screen "05_Connection_Parameters" 800x480, template "Navigation"
   on GenerateScreen: SetTag("screen_number", 5)
   ScreenModuleView "Connection_Parameters_Control_1" at 100,137 size 600x270; ScreenModuleType ""
      on Guid_{11997190-31118}: ActivateScreen("03_Connection_Control", 0)
      Guid_{11997190-30476} <- "connection_parameters"
   Rectangle "screen_background" at 0,65 size 800x415
      Appearance <- "color"
      Visibility <- "visible"
*)

(* ===== HMI "HMI_RT_1" =====
system functions are stored by id; their names below are inferred from use

ScreenModuleEditorView "Row_Wire" 400x50
   Rectangle "Border" at 0,0 size 400x50
      Appearance <- "interface.background_animate"
   IOField "IOF R0 C0" at 5,5 size 190x45; FormatPattern ????????????????????
      ProcessValue <- "text_label"
      Appearance <- "interface.cell_0_animate"
      ObjectEnable <- "interface.cell_0_enable"
      Visibility <- "interface.cell_0_visible"
   IOField "IOF R0 C1" at 200,5 size 195x45; FormatPattern 9999999
      on OnFinishInput: SetBit("interface.cell_1_input_finished")
      Visibility <- "interface.cell_1_visible"
      ObjectEnable <- "interface.cell_1_enable"
      Appearance <- "interface.cell_1_animate"
*)

(* ===== HMI "HMI_RT_1" =====
system functions are stored by id; their names below are inferred from use

ScreenModuleEditorView "Row_Wire" 400x50
   Rectangle "Border" at 0,0 size 400x50
      Appearance <- "interface.background_animate"
      Visibility <- "interface.background_visible"
   IOField "IOF R0 C0" at 5,5 size 190x45; FormatPattern ????????????????????
      Appearance <- "interface.cell_0_animate"
      ProcessValue <- "text_label"
      Visibility <- "interface.cell_0_visible"
      ObjectEnable <- "interface.cell_0_enable"
   IOField "IOF R0 C1" at 200,5 size 195x45; FormatPattern 9999999
      on OnFinishInput: SetBit("interface.cell_1_input_finished")
      Visibility <- "interface.cell_1_visible"
      Appearance <- "interface.cell_1_animate"
      ObjectEnable <- "interface.cell_1_enable"
*)

(* ===== HMI "HMI_RT_1" =====
system functions are stored by id; their names below are inferred from use

ScreenModuleEditorView "Row_Wire" 400x50
   Rectangle "Border" at 0,0 size 400x50
      Visibility <- "interface.background_visible"
      Appearance <- "interface.background_animate"
   IOField "IOF R0 C0" at 5,5 size 190x45; FormatPattern ????????????????????
      Appearance <- "interface.cell_0_animate"
      Visibility <- "interface.cell_0_visible"
      ObjectEnable <- "interface.cell_0_enable"
      ProcessValue <- "interface.cell_0_value"
   IOField "IOF R0 C1" at 200,5 size 195x45; FormatPattern 9999999
      on OnFinishInput: SetBit("interface.cell_1_input_finished")
      Visibility <- "interface.cell_1_visible"
      Appearance <- "interface.cell_1_animate"
      ObjectEnable <- "interface.cell_1_enable"
*)

(* ===== HMI "HMI_RT_1" =====
system functions are stored by id; their names below are inferred from use

ScreenModuleEditorView "Row_Wire" 400x50
   Rectangle "Border" at 0,0 size 400x50
      Visibility <- "interface.background_visible"
      Appearance <- "interface.background_animate"
   IOField "IOF R0 C0" at 5,5 size 190x45; FormatPattern ????????????????????
      Appearance <- "interface.cell_0_animate"
      Visibility <- "interface.cell_0_visible"
      ProcessValue <- "interface.cell_0_value"
      ObjectEnable <- "interface.cell_0_enable"
   IOField "IOF R0 C1" at 200,5 size 195x45; FormatPattern 9999999
      on OnFinishInput: SetBit("interface.cell_1_input_finished")
      Visibility <- "interface.cell_1_visible"
      Appearance <- "interface.cell_1_animate"
      ObjectEnable <- "interface.cell_1_enable"
*)

(* ===== HMI "HMI_RT_1" =====
system functions are stored by id; their names below are inferred from use

ScreenModuleEditorView "Row_Wire" 400x65
   Rectangle "Border" at 0,0 size 400x65
      Visibility <- "interface.background_visible"
      Appearance <- "interface.background_animate"
   TextField "TF R0 C0" at 5,5 size 190x60; Text 'Text'
      Visibility <- "interface.cell_0_visible"
   IOField "IOF R0 C1" at 200,5 size 195x60; FormatPattern 9999999
      on OnFinishInput: SetBit("interface.cell_1_input_finished")
      Visibility <- "interface.cell_1_visible"
      ObjectEnable <- "interface.cell_1_enable"
*)

(* ===== HMI "HMI_RT_1" =====
system functions are stored by id; their names below are inferred from use

ScreenModuleEditorView "Row_Wire" 600x65
   Rectangle "Border" at 0,0 size 600x65
      Visibility <- "interface.background_visible"
      Appearance <- "interface.background_animate"
   TextField "TF R0 C0" at 5,5 size 360x60; Text 'CARBON WIRE'
      Visibility <- "interface.cell_0_visible"
   IOField "IOF R0 C1" at 370,5 size 225x60; FormatPattern 9999999
      on OnFinishInput: SetBit("interface.cell_1_input_finished")
      Visibility <- "interface.cell_1_visible"
      ObjectEnable <- "interface.cell_1_enable"
*)

(* ===== HMI "HMI_RT_1" =====
system functions are stored by id; their names below are inferred from use

ScreenModuleEditorView "Row_Wire" 600x65
   Rectangle "Border" at 0,0 size 600x65
      Visibility <- "interface.background_visible"
      Appearance <- "interface.background_animate"
   TextField "TF R0 C0" at 5,5 size 360x60; Text 'CARBON WIRE'
      Visibility <- "interface.cell_0_visible"
      Appearance <- "interface.cell_0_animate"
   IOField "IOF R0 C1" at 370,5 size 225x60; FormatPattern 9999999
      on OnFinishInput: SetBit("interface.cell_1_input_finished")
      Visibility <- "interface.cell_1_visible"
      ObjectEnable <- "interface.cell_1_enable"
      Appearance <- "interface.cell_1_animate"
*)

(* ===== HMI "HMI_RT_1" =====
system functions are stored by id; their names below are inferred from use

ScreenModuleEditorView "Row_Wire_Label" 600x65
   Rectangle "Border" at 0,0 size 600x65
      Visibility <- "interface.background_visible"
      Appearance <- "interface.background_animate"
   TextField "TF R0 C0" at 5,5 size 360x60; Text 'CARBON WIRE'
      Visibility <- "interface.cell_0_visible"
      Appearance <- "interface.cell_0_animate"
   IOField "IOF R0 C1" at 370,5 size 225x60; FormatPattern 9999999
      on OnFinishInput: SetBit("interface.cell_1_input_finished")
      Visibility <- "interface.cell_1_visible"
      Appearance <- "interface.cell_1_animate"
      ObjectEnable <- "interface.cell_1_enable"
*)

(* ===== HMI "HMI_RT_1" =====

ScreenModuleEditorView "Row_Wire_Label" 600x65
   Rectangle "Border" at 0,0 size 600x65
      Visibility <- "interface.background_visible"
      Appearance <- "interface.background_animate"
   TextField "TF R0 C0" at 5,5 size 360x60; Text 'WIRE'
      Visibility <- "interface.cell_0_visible"
      Appearance <- "interface.cell_0_animate"
   TextField "TF R0 C1" at 370,5 size 225x60; Text 'LENGTH'
      Visibility <- "interface.cell_1_visible"
      Appearance <- "interface.cell_1_animate"
*)

(* ===== HMI "HMI_RT_1" =====

ScreenModuleEditorView "Divider" 600x5
   Line "line" at 10,2 size 580x0
      Appearance <- "interface.line_animate"
      Visibility <- "interface.line_visible"
   Rectangle "background" at 0,0 size 600x5
      Appearance <- "interface.background_animate"
      Visibility <- "interface.background_visible"
*)

(* ===== HMI "HMI_RT_1" =====
system functions are stored by id; their names below are inferred from use

ScreenModuleEditorView "Navigation" 800x65
   Button "Wire" at 5,5 size 390x60; TextOff 'WIRE'
      Appearance <- "interface.wire_animate"
      on Press: function_b14e0dd5("interface.wire_actuate", 0)
   Button "Material" at 400,5 size 390x60; TextOff 'MATERIAL'
      Appearance <- "interface.material_animate"
      on Press: function_b14e0dd5("interface.material_actuate", 0)
   Rectangle "Wire_Cover" at 10,60 size 380x5
      Visibility <- "interface.wire_cover_visible"
   Rectangle "Material_Cover" at 405,60 size 380x5
      Visibility <- "interface.material_cover_visible"
*)

(* ===== HMI "HMI_RT_1" =====
system functions are stored by id; their names below are inferred from use

ScreenModuleEditorView "Navigation" 800x65
   Button "Wire" at 5,5 size 390x60; TextOff 'WIRE'
      on Press: function_b14e0dd5("interface.wire_actuate", 0)
      Appearance <- "interface.wire_animate"
   Button "Material" at 400,5 size 390x60; TextOff 'MATERIAL'
      on Press: function_b14e0dd5("interface.material_actuate", 0)
      Appearance <- "interface.material_animate"
   Rectangle "Wire_Cover" at 10,60 size 380x5
      Visibility <- "interface.wire_cover_visible"
   Rectangle "Material_Cover" at 405,60 size 380x5
      Visibility <- "interface.material_cover_visible"
*)

(* ===== HMI "HMI_RT_1" =====
system functions are stored by id; their names below are inferred from use

ScreenModuleEditorView "Navigation" 800x65
   Button "Wire" at 5,5 size 392x60; TextOff 'WIRE'
      on Press: function_b14e0dd5("interface.wire_actuate", 0)
      Appearance <- "interface.wire_animate"
   Button "Material" at 402,5 size 393x60; TextOff 'MATERIAL'
      on Press: function_b14e0dd5("interface.material_actuate", 0)
      Appearance <- "interface.material_animate"
   Rectangle "Wire_Cover" at 10,60 size 382x5
      Visibility <- "interface.wire_cover_visible"
   Rectangle "Material_Cover" at 407,60 size 383x5
      Visibility <- "interface.material_cover_visible"
*)

(* ===== HMI "HMI_RT_1" =====
system functions are stored by id; their names below are inferred from use

ScreenModuleEditorView "Row_Material" 600x65
   Rectangle "Border" at 0,0 size 600x65
      Visibility <- "interface.background_visible"
      Appearance <- "interface.background_animate"
   TextField "TF R0 C0" at 5,5 size 360x60; Text 'CARBON WIRE'
      Visibility <- "interface.cell_0_visible"
      Appearance <- "interface.cell_0_animate"
   IOField "IOF R0 C1" at 370,5 size 225x60; FormatPattern 9999999
      on OnFinishInput: SetBit("interface.cell_1_input_finished")
      Visibility <- "interface.cell_1_visible"
      Appearance <- "interface.cell_1_animate"
      ObjectEnable <- "interface.cell_1_enable"
*)

(* ===== HMI "HMI_RT_1" =====
system functions are stored by id; their names below are inferred from use

ScreenModuleEditorView "Row_Material" 600x40
   Rectangle "Border" at 0,0 size 600x40
      Visibility <- "interface.background_visible"
      Appearance <- "interface.background_animate"
   IOField "IOF R0 C1" at 370,5 size 225x35; FormatPattern 9999999
      on OnFinishInput: SetBit("interface.cell_1_input_finished")
      Visibility <- "interface.cell_1_visible"
      Appearance <- "interface.cell_1_animate"
      ObjectEnable <- "interface.cell_1_enable"
   TextField "TF R0 C0" at 5,5 size 360x35; Text 'MOLYBDENUM'
      Visibility <- "interface.cell_0_visible"
      Appearance <- "interface.cell_0_animate"
*)

(* ===== HMI "HMI_RT_1" =====
system functions are stored by id; their names below are inferred from use

ScreenModuleEditorView "Row_Custom" 600x40
   Rectangle "Border" at 0,0 size 600x40
      Visibility <- "interface.background_visible"
      Appearance <- "interface.background_animate"
   IOField "IOF R0 C1" at 370,5 size 225x35; FormatPattern 9999999
      on OnFinishInput: SetBit("interface.cell_1_input_finished")
      Visibility <- "interface.cell_1_visible"
      Appearance <- "interface.cell_1_animate"
      ObjectEnable <- "interface.cell_1_enable"
   TextField "TF R0 C0" at 5,5 size 360x35; Text 'MOLYBDENUM'
      Visibility <- "interface.cell_0_visible"
      Appearance <- "interface.cell_0_animate"
*)

(* ===== HMI "HMI_RT_1" =====
system functions are stored by id; their names below are inferred from use

ScreenModuleEditorView "Row_Custom" 600x40
   Rectangle "Border" at 0,0 size 600x40
      Visibility <- "interface.background_visible"
      Appearance <- "interface.background_animate"
   IOField "IOF R0 C0" at 5,5 size 360x35; FormatPattern ???????????????
      on OnFinishInput: SetBit("interface.cell_0_input_finished")
      Appearance <- "interface.cell_0_animate"
      ObjectEnable <- "interface.cell_0_enable"
      Visibility <- "interface.cell_0_visible"
   IOField "IOF R0 C1" at 370,5 size 225x35; FormatPattern 9999999
      on OnFinishInput: SetBit("interface.cell_1_input_finished")
      Visibility <- "interface.cell_1_visible"
      Appearance <- "interface.cell_1_animate"
      ObjectEnable <- "interface.cell_1_enable"
*)

(* ===== HMI "HMI_RT_1" =====
system functions are stored by id; their names below are inferred from use

ScreenModuleEditorView "Row_Material_Label" 600x40
   Rectangle "Border" at 0,0 size 600x40
      Visibility <- "interface.background_visible"
      Appearance <- "interface.background_animate"
   IOField "IOF R0 C1" at 370,5 size 225x35; FormatPattern 9999999
      on OnFinishInput: SetBit("interface.cell_1_input_finished")
      Visibility <- "interface.cell_1_visible"
      Appearance <- "interface.cell_1_animate"
      ObjectEnable <- "interface.cell_1_enable"
   TextField "TF R0 C0" at 5,5 size 360x35; Text 'MOLYBDENUM'
      Visibility <- "interface.cell_0_visible"
      Appearance <- "interface.cell_0_animate"
*)

(* ===== HMI "HMI_RT_1" =====

ScreenModuleEditorView "Row_Material_Label" 600x40
   Rectangle "Border" at 0,0 size 600x40
      Visibility <- "interface.background_visible"
      Appearance <- "interface.background_animate"
   TextField "TF R0 C0" at 5,5 size 360x35; Text 'MATERIAL'
      Visibility <- "interface.cell_0_visible"
      Appearance <- "interface.cell_0_animate"
   TextField "TF R0 C1" at 370,5 size 225x35; Text 'BAGS'
      Appearance <- "interface.cell_1_animate"
      Visibility <- "interface.cell_1_visible"
*)

(* ===== HMI "HMI_RT_1" =====
system functions are stored by id; their names below are inferred from use

ScreenModuleEditorView "Row_Wire" 600x65
   Rectangle "Border" at 0,0 size 600x65
      Visibility <- "interface.background_visible"
   TextField "TF R0 C0" at 5,5 size 360x60; Text 'CARBON WIRE'
      Visibility <- "interface.cell_0_visible"
   IOField "IOF R0 C1" at 370,5 size 225x60; FormatPattern 9999999
      on OnFinishInput: SetBit("interface.cell_1_input_finished")
      Visibility <- "interface.cell_1_visible"
      Appearance <- "interface.cell_1_animate"
      ObjectEnable <- "interface.cell_1_enable"
      on Activate: SetBit("interface.cell_1_active")
      on Deactivate: ResetBit("interface.cell_1_active")
*)

(* ===== HMI "HMI_RT_1" =====

ScreenModuleEditorView "Divider" 600x5
   Line "line" at 10,2 size 580x0
      Visibility <- "interface.line_visible"
      Appearance <- "interface.line_animate"
   Rectangle "background" at 0,0 size 600x5
      Visibility <- "interface.background_visible"
      Appearance <- "interface.background_animate"
*)

(* ===== HMI "HMI_RT_1" =====
system functions are stored by id; their names below are inferred from use

ScreenModuleEditorView "Row_Material" 600x40
   Rectangle "Border" at 0,0 size 600x40
      Visibility <- "interface.background_visible"
      Appearance <- "interface.background_animate"
   IOField "IOF R0 C1" at 370,5 size 225x35; FormatPattern 9999999
      on OnFinishInput: SetBit("interface.cell_1_input_finished")
      Visibility <- "interface.cell_1_visible"
      Appearance <- "interface.cell_1_animate"
      ObjectEnable <- "interface.cell_1_enable"
   TextField "TF R0 C0" at 5,5 size 360x35; Text 'MOLYBDENUM'
      Visibility <- "interface.cell_0_visible"
      Appearance <- "interface.cell_0_animate"
*)

(* ===== HMI "HMI_RT_1" =====
system functions are stored by id; their names below are inferred from use

ScreenModuleEditorView "Navigation" 800x65
   Button "Wire" at 5,5 size 392x60; TextOff 'WIRE'
      on Press: function_b14e0dd5("interface.wire_actuate", 0)
      Appearance <- "interface.wire_animate"
      ObjectEnable <- "interface.wire_enable"
      Visibility <- "interface.wire_visible"
   Button "Material" at 402,5 size 393x60; TextOff 'MATERIAL'
      on Press: function_b14e0dd5("interface.material_actuate", 0)
      Appearance <- "interface.material_animate"
      ObjectEnable <- "interface.material_enable"
      Visibility <- "interface.material_visible"
   Rectangle "Background" at 0,0 size 800x65
      Appearance <- "interface.background_animate"
      Visibility <- "interface.background_visible"
   Rectangle "Wire_Cover" at 10,60 size 382x5
      Visibility <- "interface.wire_cover_visible"
      Appearance <- "interface.wire_cover_animate"
   Rectangle "Material_Cover" at 407,60 size 383x5
      Visibility <- "interface.material_cover_visible"
      Appearance <- "interface.material_cover_animate"
   Line "Bottom_Line" at 0,62 size 800x0
      Appearance <- "interface.bottom_line_animate"
      Visibility <- "interface.bottom_line_visible"
*)

(* ===== HMI "HMI_RT_1" =====
system functions are stored by id; their names below are inferred from use

ScreenModuleEditorView "Navigation" 800x65
   Button "Wire" at 5,5 size 392x60; TextOff 'WIRE'
      on Press: function_b14e0dd5("interface.wire_actuate", 0)
      Appearance <- "interface.wire_animate"
      ObjectEnable <- "interface.wire_enable"
      Visibility <- "interface.wire_visible"
   Button "Material" at 402,5 size 393x60; TextOff 'MATERIAL'
      on Press: function_b14e0dd5("interface.material_actuate", 0)
      Appearance <- "interface.material_animate"
      ObjectEnable <- "interface.material_enable"
      Visibility <- "interface.material_visible"
   Rectangle "Background" at 0,0 size 800x65
      Visibility <- "interface.background_visible"
      Appearance <- "interface.background_animate"
   Rectangle "Wire_Cover" at 10,60 size 382x5
      Visibility <- "interface.wire_cover_visible"
      Appearance <- "interface.wire_cover_animate"
   Rectangle "Material_Cover" at 407,60 size 383x5
      Visibility <- "interface.material_cover_visible"
      Appearance <- "interface.material_cover_animate"
   Line "Bottom_Line" at 0,62 size 800x0
      Visibility <- "interface.bottom_line_visible"
      Appearance <- "interface.bottom_line_animate"
*)

(* ===== HMI "HMI_RT_1" =====
system functions are stored by id; their names below are inferred from use

ScreenModuleEditorView "Navigation" 800x65
   Button "Wire" at 5,5 size 392x60; TextOff 'WIRE'
      on Press: function_b14e0dd5("interface.wire_actuate", 0)
      Appearance <- "interface.wire_animate"
      ObjectEnable <- "interface.wire_enable"
      Visibility <- "interface.wire_visible"
   Button "Material" at 402,5 size 393x60; TextOff 'MATERIAL'
      on Press: function_b14e0dd5("interface.material_actuate", 0)
      Appearance <- "interface.material_animate"
      ObjectEnable <- "interface.material_enable"
      Visibility <- "interface.material_visible"
   Rectangle "Background" at 0,0 size 800x65
      Visibility <- "interface.background_visible"
      Appearance <- "interface.background_animate"
   Rectangle "Wire_Cover" at 10,60 size 382x5
      Visibility <- "interface.wire_cover_visible"
      Appearance <- "interface.wire_cover_animate"
   Rectangle "Material_Cover" at 407,60 size 383x5
      Visibility <- "interface.material_cover_visible"
      Appearance <- "interface.material_cover_animate"
   Line "Bottom_Line" at 0,62 size 800x0
      Visibility <- "interface.bottom_line_visible"
      Appearance <- "interface.bottom_line_animate"
*)

(* ===== HMI "HMI_RT_1" =====
system functions are stored by id; their names below are inferred from use

ScreenModuleEditorView "Navigation" 800x65
   Button "Wire" at 5,5 size 392x60; TextOff 'WIRE'
      on Press: function_b14e0dd5("interface.wire_actuate", 0)
      Appearance <- "interface.wire_animate"
      ObjectEnable <- "interface.wire_enable"
      Visibility <- "interface.wire_visible"
   Button "Material" at 402,5 size 393x60; TextOff 'MATERIAL'
      on Press: function_b14e0dd5("interface.material_actuate", 0)
      Appearance <- "interface.material_animate"
      ObjectEnable <- "interface.material_enable"
      Visibility <- "interface.material_visible"
   Rectangle "Background" at 0,0 size 800x65
      Visibility <- "interface.background_visible"
      Appearance <- "interface.background_animate"
   Rectangle "Wire_Cover" at 10,60 size 382x5
      Visibility <- "interface.wire_cover_visible"
      Appearance <- "interface.wire_cover_animate"
   Rectangle "Material_Cover" at 407,60 size 383x5
      Visibility <- "interface.material_cover_visible"
      Appearance <- "interface.material_cover_animate"
   Line "Bottom_Line" at 0,62 size 800x0
      Visibility <- "interface.bottom_line_visible"
      Appearance <- "interface.bottom_line_animate"
*)

(* ===== HMI "HMI_RT_1" =====
system functions are stored by id; their names below are inferred from use

ScreenModuleEditorView "Navigation" 800x65
   Button "wire_button" at 5,5 size 260x60; TextOff 'WIRE'
      on Press: function_b14e0dd5("interface.wire_actuate", 0)
      Appearance <- "interface.wire_animate"
      ObjectEnable <- "interface.wire_enable"
      Visibility <- "interface.wire_visible"
   Button "material_button" at 270,5 size 260x60; TextOff 'MATERIAL'
      on Press: function_b14e0dd5("interface.material_actuate", 0)
      Appearance <- "interface.material_animate"
      ObjectEnable <- "interface.material_enable"
      Visibility <- "interface.material_visible"
   Button "communications_status_button" at 535,5 size 260x60; TextOff 'COMMUNICATIONS STATUS'
      on Press: function_b14e0dd5("interface.communications_status_actuate", 0)
      Visibility <- "interface.communications_status_visible"
      ObjectEnable <- "interface.communications_status_enable"
      Appearance <- "interface.communications_status_animate"
   Rectangle "Background" at 0,0 size 800x65
      Visibility <- "interface.background_visible"
      Appearance <- "interface.background_animate"
   Rectangle "wire_cover" at 10,60 size 250x5
      Visibility <- "interface.wire_cover_visible"
      Appearance <- "interface.wire_cover_animate"
   Rectangle "material_cover" at 275,60 size 250x5
      Visibility <- "interface.material_cover_visible"
      Appearance <- "interface.material_cover_animate"
   Rectangle "communications_status_cover" at 540,60 size 250x5
      Appearance <- "interface.communications_status_cover_animate"
      Visibility <- "interface.communications_status_cover_visible"
   Line "Bottom_Line" at 0,62 size 800x0
      Visibility <- "interface.bottom_line_visible"
      Appearance <- "interface.bottom_line_animate"
*)

(* ===== HMI "HMI_RT_1" =====

ScreenModuleEditorView "Row_Wire_Label" 600x65
   Rectangle "Border" at 0,0 size 600x65
      Visibility <- "interface.background_visible"
      Appearance <- "interface.background_animate"
   TextField "TF R0 C0" at 5,5 size 360x60; Text 'WIRE'
      Visibility <- "interface.cell_0_visible"
      Appearance <- "interface.cell_0_animate"
   TextField "TF R0 C1" at 370,5 size 225x60; Text 'LENGTH'
      Visibility <- "interface.cell_1_visible"
      Appearance <- "interface.cell_1_animate"
*)

(* ===== HMI "HMI_RT_1" =====
system functions are stored by id; their names below are inferred from use

ScreenModuleEditorView "Row_Wire" 600x65
   Rectangle "Border" at 0,0 size 600x65
      Visibility <- "interface.background_visible"
      Appearance <- "interface.background_animate"
   TextField "TF R0 C0" at 5,5 size 360x60; Text 'CARBON WIRE'
      Visibility <- "interface.cell_0_visible"
      Appearance <- "interface.cell_0_animate"
   IOField "IOF R0 C1" at 370,5 size 225x60; FormatPattern 9999999
      on OnFinishInput: SetBit("interface.cell_1_input_finished")
      on Deactivate: ResetBit("interface.cell_1_active")
      on Activate: SetBit("interface.cell_1_active")
      Visibility <- "interface.cell_1_visible"
      ObjectEnable <- "interface.cell_1_enable"
      Appearance <- "interface.cell_1_animate"
*)

(* ===== HMI "HMI_RT_1" =====

ScreenModuleEditorView "Row_Wire_Label" 600x65
   Rectangle "Border" at 0,0 size 600x65
      Visibility <- "interface.background_visible"
      Appearance <- "interface.background_animate"
   TextField "TF R0 C0" at 5,5 size 360x60; Text 'WIRE'
      Visibility <- "interface.cell_0_visible"
      Appearance <- "interface.cell_0_animate"
   TextField "TF R0 C1" at 370,5 size 225x60; Text 'LENGTH'
      Visibility <- "interface.cell_1_visible"
      Appearance <- "interface.cell_1_animate"
*)

(* ===== HMI "HMI_RT_1" =====
system functions are stored by id; their names below are inferred from use

ScreenModuleEditorView "Row_Material" 600x40
   Rectangle "Border" at 0,0 size 600x40
      Visibility <- "interface.background_visible"
      Appearance <- "interface.background_animate"
   TextField "TF R0 C0" at 5,5 size 360x35; Text 'MOLYBDENUM'
      Visibility <- "interface.cell_0_visible"
      Appearance <- "interface.cell_0_animate"
   IOField "IOF R0 C1" at 370,5 size 225x35; FormatPattern 9999999
      on OnFinishInput: SetBit("interface.cell_1_input_finished")
      Visibility <- "interface.cell_1_visible"
      ObjectEnable <- "interface.cell_1_enable"
      Appearance <- "interface.cell_1_animate"
      on Activate: SetBit("interface.cell_1_active")
      on Deactivate: ResetBit("interface.cell_1_active")
*)

(* ===== HMI "HMI_RT_1" =====

ScreenModuleEditorView "Row_Material_Label" 600x40
   Rectangle "Border" at 0,0 size 600x40
      Visibility <- "interface.background_visible"
      Appearance <- "interface.background_animate"
   TextField "TF R0 C0" at 5,5 size 360x35; Text 'MATERIAL'
      Visibility <- "interface.cell_0_visible"
      Appearance <- "interface.cell_0_animate"
   TextField "TF R0 C1" at 370,5 size 225x35; Text 'BAGS'
      Visibility <- "interface.cell_1_visible"
      Appearance <- "interface.cell_1_animate"
*)

(* ===== HMI "HMI_RT_1" =====
system functions are stored by id; their names below are inferred from use

ScreenModuleEditorView "Row_Custom" 600x40
   Rectangle "Border" at 0,0 size 600x40
      Visibility <- "interface.background_visible"
      Appearance <- "interface.background_animate"
   IOField "IOF R0 C0" at 5,5 size 360x35; FormatPattern ???????????????
      on OnFinishInput: SetBit("interface.cell_0_input_finished")
      ObjectEnable <- "interface.cell_0_enable"
      Visibility <- "interface.cell_0_visible"
      Appearance <- "interface.cell_0_animate"
      on Activate: SetBit("interface.cell_0_activate")
      on Deactivate: ResetBit("interface.cell_0_activate")
   IOField "IOF R0 C1" at 370,5 size 225x35; FormatPattern 9999999
      on OnFinishInput: SetBit("interface.cell_1_input_finished")
      Visibility <- "interface.cell_1_visible"
      ObjectEnable <- "interface.cell_1_enable"
      Appearance <- "interface.cell_0_animate"
      on Activate: SetBit("interface.cell_1_activate")
      on Deactivate: ResetBit("interface.cell_1_activate")
*)

(* ===== HMI "HMI_RT_1" =====
system functions are stored by id; their names below are inferred from use

ScreenModuleEditorView "Row_Wire" 600x65
   Rectangle "Border" at 0,0 size 600x65
      Visibility <- "interface.background_visible"
      Appearance <- "interface.background_animate"
   TextField "TF R0 C0" at 5,5 size 360x60; Text 'CARBON WIRE'
      Visibility <- "interface.cell_0_visible"
      Appearance <- "interface.cell_0_animate"
   IOField "IOF R0 C1" at 370,5 size 225x60; FormatPattern ???????
      on Deactivate: ResetBit("interface.cell_1_active")
      on OnFinishInput: SetBit("interface.cell_1_input_finished")
      on Activate: SetBit("interface.cell_1_active")
      Visibility <- "interface.cell_1_visible"
      ObjectEnable <- "interface.cell_1_enable"
      Appearance <- "interface.cell_1_animate"
      ProcessValue <- "interface.cell_1_value"
*)

(* ===== HMI "HMI_RT_1" =====
system functions are stored by id; their names below are inferred from use

ScreenModuleEditorView "Row_Material" 600x40
   Rectangle "Border" at 0,0 size 600x40
      Visibility <- "interface.background_visible"
      Appearance <- "interface.background_animate"
   TextField "TF R0 C0" at 5,5 size 360x35; Text 'MOLYBDENUM'
      Visibility <- "interface.cell_0_visible"
      Appearance <- "interface.cell_0_animate"
   IOField "IOF R0 C1" at 370,5 size 225x35; FormatPattern ?????????
      on OnFinishInput: SetBit("interface.cell_1_input_finished")
      on Deactivate: ResetBit("interface.cell_1_active")
      on Activate: SetBit("interface.cell_1_active")
      Appearance <- "interface.cell_1_animate"
      Visibility <- "interface.cell_1_visible"
      ObjectEnable <- "interface.cell_1_enable"
      ProcessValue <- "interface.cell_1_value"
*)

(* ===== HMI "HMI_RT_1" =====
system functions are stored by id; their names below are inferred from use

ScreenModuleEditorView "Row_Custom" 600x40
   Rectangle "Border" at 0,0 size 600x40
      Visibility <- "interface.background_visible"
      Appearance <- "interface.background_animate"
   IOField "IOF R0 C0" at 5,5 size 360x35; FormatPattern ???????????????
      on OnFinishInput: SetBit("interface.cell_0_input_finished")
      on Deactivate: ResetBit("interface.cell_0_activate")
      on Activate: SetBit("interface.cell_0_activate")
      Appearance <- "interface.cell_0_animate"
      Visibility <- "interface.cell_0_visible"
      ObjectEnable <- "interface.cell_0_enable"
      ProcessValue <- "interface.cell_0_value"
   IOField "IOF R0 C1" at 370,5 size 225x35; FormatPattern ?????????
      on OnFinishInput: SetBit("interface.cell_1_input_finished")
      on Deactivate: ResetBit("interface.cell_1_activate")
      on Activate: SetBit("interface.cell_1_activate")
      Appearance <- "interface.cell_0_animate"
      Visibility <- "interface.cell_1_visible"
      ObjectEnable <- "interface.cell_1_enable"
      ProcessValue <- "interface.cell_1_value"
*)

(* ===== HMI "HMI_RT_1" =====
system functions are stored by id; their names below are inferred from use

ScreenModuleEditorView "Row_Custom" 600x40
   Rectangle "Border" at 0,0 size 600x40
      Visibility <- "interface.background_visible"
      Appearance <- "interface.background_animate"
   IOField "IOF R0 C0" at 5,5 size 360x35; FormatPattern ???????????????
      on Deactivate: ResetBit("interface.cell_0_activate")
      on OnFinishInput: SetBit("interface.cell_0_input_finished")
      on Activate: SetBit("interface.cell_0_activate")
      ProcessValue <- "interface.cell_0_value"
      Visibility <- "interface.cell_0_visible"
      Appearance <- "interface.cell_0_animate"
      ObjectEnable <- "interface.cell_0_enable"
   IOField "IOF R0 C1" at 370,5 size 225x35; FormatPattern ?????????
      on Deactivate: ResetBit("interface.cell_1_activate")
      on OnFinishInput: SetBit("interface.cell_1_input_finished")
      on Activate: SetBit("interface.cell_1_activate")
      ProcessValue <- "interface.cell_1_value"
      Visibility <- "interface.cell_1_visible"
      ObjectEnable <- "interface.cell_1_enable"
      Appearance <- "interface.cell_1_animate"
*)

(* ===== HMI "HMI_RT_1" =====

text list "Send Code Descriptions Short": 0 'SEND SUCCESSFUL'; 28672 'NO JOB'; 28673 'DATA ACCESSED DURING JOB'; 28674 'JOB PROCESSING'; 32901 'MAX LENGTH EXCEEDED'; 32902 'INVALID ID OUT OF RANGE'; 32904 'LENGTH EXCEEDS DATA RANGE'; 32929 'NO CONNECTION'; 32947 'UDP CONNECTION'; 32963 'CONNECTION BUSY'; 32964 'REQUEST DURING PARAM ASSIGNMENT'; 32965 'PARTNER TERMINATED CONNECTION'; 32966 'PARTNER UNAVAILABLE'; 32967 'TIMEOUT'; 65535 'NOT CALLED'

text list "Connect Code Descriptions Short": 0 'CONNECTION SUCCESSFUL'; 28672 'NO JOB'; 28673 'START JOB'; 28674 'PROCESSING JOB'; 32901 'ID INVALID: ALREADY IN USE'; 32902 'ID INVALID: OUT OF RANGE'; 32903 'MAX CONNECTIONS REACHED'; 32905 'NO CONNECTION DATA STORED'; 32922 'INVALID CONNECTION DATA'; 32923 'NO CONNECTION HARDWARE'; 32928 'GROUP ERROR'; 32929 'LOCAL PORT IN USE'; 32930 'REMOTE PORT IN USE'; 32931 'CONNECTION ALREADY ESTABLISHED'; 32932 'INVALID IP ADDRESS'; 32933 'DUPLICATE CONNECTION ID'; 32935 'DICONNECT REQUEST WHILE CONNECTING'; 32946 'CONNECT DATA IN LOAD MEMORY'; 32948 'ISO ON TCP VIOLATION'; 32949 'NON PASSIVE UDP CONNECTION REQUEST'; 32950 'INVALID CONNECTION TYPE'; 32951 'CONNECTION PARAMETER ERROR'; 32952 'DATA/PARAMETER MISMATCH'; 32963 'MAX CONNECTIONS EXCEEDED'; 32964 'FIREWALL'; 65535 'STATE: DISCONNECT'; 32966 'PARTNER UNAVAILABLE'

text list "Disconnect Code Descriptions Short": 0 'DISCONNECTION SUCCESSFUL'; 28672 'NO JOB'; 28673 'JOB STARTED'; 28674 'REQUEST DURING EXECUTION'; 32902 'ID INVALID: OUT OF RANGE'; 32931 'CONNECTION ALREADY TERMINATED'; 32964 'REQUEST DURING PARAM ASSIGNMENT'; 65535 'STATE: CONNECT'

text list "Text List Select": 0 ''; 1 ''; 2 ''; 3 ''

ScreenModuleEditorView "Connection_Status_Element" 392x110
   TextField "operation_label" at 0,0 size 110x110; Text 'S'
      Visibility <- "interface.operation_label_visible"
      Appearance <- "interface.operation_label_animate"
   TextField "done_status_indicator" at 110,0 size 94x27; Text 'DONE'
      Appearance <- "interface.done_status_indicator_animate"
      Visibility <- "interface.done_status_indicator_visible"
   TextField "busy_status_indicator" at 204,0 size 94x27; Text 'BUSY'
      Visibility <- "interface.busy_status_indicator_visible"
      Appearance <- "interface.busy_status_indicator_animate"
   TextField "error_status_indicator" at 298,0 size 94x27; Text 'ERROR'
      Appearance <- "interface.error_status_indicator_animate"
      Visibility <- "interface.error_status_indicator_visible"
   TextField "status_code_label" at 110,27 size 82x28; Text 'CODE:'
      Visibility <- "interface.status_code_label_visible"
      Appearance <- "interface.status_code_label_animate"
   IOField "status_code" at 192,27 size 200x28; FormatPattern ??????
      Visibility <- "interface.status_code_value_visible"
      Appearance <- "interface.status_code_value_animate"
      ProcessValue <- "interface.status_code_value"
   SymbolicIOField "status_description" at 110,55 size 282x55; TextOn '1'; TextOff '0'; TextList "Text List Select"
      ProcessValue <- "operation_list_selector"
      Appearance <- "interface.status_code_description_animate"
      Visibility <- "interface.status_code_description_visible"
*)

(* ===== HMI "HMI_RT_1" =====

ScreenModuleEditorView "Connection_Status_Header" 392x55
   TextField "header" at 0,0 size 392x55; Text '[PARTNER NAME] COMMUNICATIONS'
      Appearance <- "interface.animate"
      Visibility <- "interface.visible"
*)

(* ===== HMI "HMI_RT_1" =====

ScreenModuleEditorView "Connection_Status_Header" 392x55
   TextField "header" at 0,0 size 392x55; Text '[PARTNER NAME] COMMUNICATIONS'
      Visibility <- "interface.visible"
      Appearance <- "interface.animate"
*)

(* ===== HMI "HMI_RT_1" =====
system functions are stored by id; their names below are inferred from use

text list "Send Code Descriptions Short": 0 'SEND SUCCESSFUL'; 28672 'NO JOB'; 28673 'DATA ACCESSED DURING JOB'; 28674 'JOB PROCESSING'; 32901 'MAX LENGTH EXCEEDED'; 32902 'INVALID ID OUT OF RANGE'; 32904 'LENGTH EXCEEDS DATA RANGE'; 32929 'NO CONNECTION'; 32947 'UDP CONNECTION'; 32963 'CONNECTION BUSY'; 32964 'REQUEST DURING PARAM ASSIGNMENT'; 32965 'PARTNER TERMINATED CONNECTION'; 32966 'PARTNER UNAVAILABLE'; 32967 'TIMEOUT'; 65535 'NOT CALLED'

text list "Connect Code Descriptions Short": 0 'CONNECTION SUCCESSFUL'; 28672 'NO JOB'; 28673 'START JOB'; 28674 'PROCESSING JOB'; 32901 'ID INVALID: ALREADY IN USE'; 32902 'ID INVALID: OUT OF RANGE'; 32903 'MAX CONNECTIONS REACHED'; 32905 'NO CONNECTION DATA STORED'; 32922 'INVALID CONNECTION DATA'; 32923 'NO CONNECTION HARDWARE'; 32928 'GROUP ERROR'; 32929 'LOCAL PORT IN USE'; 32930 'REMOTE PORT IN USE'; 32931 'CONNECTION ALREADY ESTABLISHED'; 32932 'INVALID IP ADDRESS'; 32933 'DUPLICATE CONNECTION ID'; 32935 'DICONNECT REQUEST WHILE CONNECTING'; 32946 'CONNECT DATA IN LOAD MEMORY'; 32948 'ISO ON TCP VIOLATION'; 32949 'NON PASSIVE UDP CONNECTION REQUEST'; 32950 'INVALID CONNECTION TYPE'; 32951 'CONNECTION PARAMETER ERROR'; 32952 'DATA/PARAMETER MISMATCH'; 32963 'MAX CONNECTIONS EXCEEDED'; 32964 'FIREWALL'; 65535 'STATE: DISCONNECT'; 32966 'PARTNER UNAVAILABLE'

text list "Disconnect Code Descriptions Short": 0 'DISCONNECTION SUCCESSFUL'; 28672 'NO JOB'; 28673 'JOB STARTED'; 28674 'REQUEST DURING EXECUTION'; 32902 'ID INVALID: OUT OF RANGE'; 32931 'CONNECTION ALREADY TERMINATED'; 32964 'REQUEST DURING PARAM ASSIGNMENT'; 65535 'STATE: CONNECT'

text list "Text List Select": 0 ''; 1 ''; 2 ''; 3 ''

ScreenModuleEditorView "Connection_Status_Element" 392x110
   TextField "operation_label" at 0,0 size 110x110; Text 'S'
      Visibility <- "interface.operation_label_visible"
      Appearance <- "interface.operation_label_animate"
   TextField "done_status_indicator" at 110,0 size 94x27; Text 'DONE'
      Visibility <- "interface.done_status_indicator_visible"
      Appearance <- "interface.done_status_indicator_animate"
   TextField "busy_status_indicator" at 204,0 size 94x27; Text 'BUSY'
      Visibility <- "interface.busy_status_indicator_visible"
      Appearance <- "interface.busy_status_indicator_animate"
   TextField "error_status_indicator" at 298,0 size 94x27; Text 'ERROR'
      Visibility <- "interface.error_status_indicator_visible"
      Appearance <- "interface.error_status_indicator_animate"
   TextField "status_code_label" at 110,27 size 82x28; Text 'CODE:'
      Visibility <- "interface.status_code_label_visible"
      Appearance <- "interface.status_code_label_animate"
   IOField "status_code" at 192,27 size 200x28; FormatPattern ??????
      Appearance <- "interface.status_code_value_animate"
      Visibility <- "interface.status_code_value_visible"
      ProcessValue <- "interface.status_code_value"
   SymbolicIOField "status_description" at 110,55 size 282x55; TextOn '1'; TextOff '0'; TextList "Text List Select"
      Appearance <- "interface.status_code_description_animate"
      ProcessValue <- "operation_list_selector"
      Visibility <- "interface.status_code_description_visible"
   Button "operation_left" at 0,0 size 110x110; TextOff 'Text'
      on Press: function_b14e0dd5("interface.operation_button_actuate", 0)
      ObjectEnable <- "interface.operation_button_enable"
      Visibility <- "interface.operation_button_visible"
   Button "operation_top" at 110,0 size 282x55; TextOff 'Text'
      ObjectEnable <- "interface.operation_button_actuate"
      Visibility <- "interface.operation_button_visible"
      on Press: function_b14e0dd5("interface.operation_button_actuate", 0)
   Button "show_status" at 110,55 size 282x55; TextOff 'Text'
      ObjectEnable <- "interface.show_status_code_description_button_enable"
      Visibility <- "interface.show_status_code_description_button_visible"
      on Press: function_b14e0dd5("interface.show_status_code_description_button_actuate", 0)
*)

(* ===== HMI "HMI_RT_1" =====
system functions are stored by id; their names below are inferred from use

ScreenModuleEditorView "Navigation" 800x65
   Button "wire_button" at 5,5 size 260x60; TextOff 'WIRE'
      on Press: function_b14e0dd5("interface.wire_actuate", 0)
      Appearance <- "interface.wire_animate"
      ObjectEnable <- "interface.wire_enable"
      Visibility <- "interface.wire_visible"
   Button "material_button" at 270,5 size 260x60; TextOff 'MATERIAL'
      on Press: function_b14e0dd5("interface.material_actuate", 0)
      Appearance <- "interface.material_animate"
      ObjectEnable <- "interface.material_enable"
      Visibility <- "interface.material_visible"
   Button "communications_status_button" at 535,5 size 260x60; TextOff 'CONNECTIONS'
      on Press: function_b14e0dd5("interface.communications_status_actuate", 0)
      Visibility <- "interface.communications_status_visible"
      ObjectEnable <- "interface.communications_status_enable"
      Appearance <- "interface.communications_status_animate"
   Rectangle "Background" at 0,0 size 800x65
      Visibility <- "interface.background_visible"
      Appearance <- "interface.background_animate"
   Rectangle "wire_cover" at 10,60 size 250x5
      Visibility <- "interface.wire_cover_visible"
      Appearance <- "interface.wire_cover_animate"
   Rectangle "material_cover" at 275,60 size 250x5
      Visibility <- "interface.material_cover_visible"
      Appearance <- "interface.material_cover_animate"
   Rectangle "communications_status_cover" at 540,60 size 250x5
      Visibility <- "interface.communications_status_cover_visible"
      Appearance <- "interface.communications_status_cover_animate"
   Line "Bottom_Line" at 0,62 size 800x0
      Visibility <- "interface.bottom_line_visible"
      Appearance <- "interface.bottom_line_animate"
*)

(* ===== HMI "HMI_RT_1" =====
system functions are stored by id; their names below are inferred from use

text list "Send Code Descriptions Short": 0 'SEND SUCCESSFUL'; 28672 'NO JOB'; 28673 'DATA ACCESSED DURING JOB'; 28674 'JOB PROCESSING'; 32901 'MAX LENGTH EXCEEDED'; 32902 'INVALID ID OUT OF RANGE'; 32904 'LENGTH EXCEEDS DATA RANGE'; 32929 'NO CONNECTION'; 32947 'UDP CONNECTION'; 32963 'CONNECTION BUSY'; 32964 'REQUEST DURING PARAM ASSIGNMENT'; 32965 'PARTNER TERMINATED CONNECTION'; 32966 'PARTNER UNAVAILABLE'; 32967 'TIMEOUT'; 65535 'NOT CALLED'

text list "Connect Code Descriptions Short": 0 'CONNECTION SUCCESSFUL'; 28672 'NO JOB'; 28673 'START JOB'; 28674 'PROCESSING JOB'; 32901 'ID INVALID: ALREADY IN USE'; 32902 'ID INVALID: OUT OF RANGE'; 32903 'MAX CONNECTIONS REACHED'; 32905 'NO CONNECTION DATA STORED'; 32922 'INVALID CONNECTION DATA'; 32923 'NO CONNECTION HARDWARE'; 32928 'GROUP ERROR'; 32929 'LOCAL PORT IN USE'; 32930 'REMOTE PORT IN USE'; 32931 'CONNECTION ALREADY ESTABLISHED'; 32932 'INVALID IP ADDRESS'; 32933 'DUPLICATE CONNECTION ID'; 32935 'DICONNECT REQUEST WHILE CONNECTING'; 32946 'CONNECT DATA IN LOAD MEMORY'; 32948 'ISO ON TCP VIOLATION'; 32949 'NON PASSIVE UDP CONNECTION REQUEST'; 32950 'INVALID CONNECTION TYPE'; 32951 'CONNECTION PARAMETER ERROR'; 32952 'DATA/PARAMETER MISMATCH'; 32963 'MAX CONNECTIONS EXCEEDED'; 32964 'FIREWALL'; 65535 'STATE: DISCONNECT'; 32966 'PARTNER UNAVAILABLE'

text list "Disconnect Code Descriptions Short": 0 'DISCONNECTION SUCCESSFUL'; 28672 'NO JOB'; 28673 'JOB STARTED'; 28674 'REQUEST DURING EXECUTION'; 32902 'ID INVALID: OUT OF RANGE'; 32931 'CONNECTION ALREADY TERMINATED'; 32964 'REQUEST DURING PARAM ASSIGNMENT'; 65535 'STATE: CONNECT'

text list "Text List Select": 0 ''; 1 ''; 2 ''; 3 ''

ScreenModuleEditorView "Connection_Status_Element" 392x110
   TextField "operation_label" at 0,0 size 110x110; Text 'S'
      Visibility <- "interface.operation_label_visible"
      Appearance <- "interface.operation_label_animate"
   TextField "done_status_indicator" at 110,0 size 94x27; Text 'DONE'
      Visibility <- "interface.done_status_indicator_visible"
      Appearance <- "interface.done_status_indicator_animate"
   TextField "busy_status_indicator" at 204,0 size 94x27; Text 'BUSY'
      Visibility <- "interface.busy_status_indicator_visible"
      Appearance <- "interface.busy_status_indicator_animate"
   TextField "error_status_indicator" at 298,0 size 94x27; Text 'ERROR'
      Visibility <- "interface.error_status_indicator_visible"
      Appearance <- "interface.error_status_indicator_animate"
   TextField "status_code_label" at 110,27 size 82x28; Text 'CODE:'
      Visibility <- "interface.status_code_label_visible"
      Appearance <- "interface.status_code_label_animate"
   IOField "status_code" at 192,27 size 200x28; FormatPattern ??????
      Appearance <- "interface.status_code_value_animate"
      Visibility <- "interface.status_code_value_visible"
      ProcessValue <- "interface.status_code_value"
   SymbolicIOField "status_description" at 110,55 size 282x55; TextOn '1'; TextOff '0'; TextList "Text List Select"
      Appearance <- "interface.status_code_description_animate"
      ProcessValue <- "operation_list_selector"
      Visibility <- "interface.status_code_description_visible"
   Button "operation_left" at 0,0 size 110x110; TextOff 'Text'
      on Press: function_b14e0dd5("interface.operation_button_actuate", 0)
      Visibility <- "interface.operation_button_visible"
      ObjectEnable <- "interface.operation_button_enable"
   Button "operation_top" at 110,0 size 282x55; TextOff 'Text'
      on Press: function_b14e0dd5("interface.operation_button_actuate", 0)
      Visibility <- "interface.operation_button_visible"
      ObjectEnable <- "interface.operation_button_actuate"
   Button "show_status" at 110,55 size 282x55; TextOff 'Text'
      on Press: function_b14e0dd5("interface.show_status_code_description_button_actuate", 0)
      Visibility <- "interface.show_status_code_description_button_visible"
      ObjectEnable <- "interface.show_status_code_description_button_enable"
*)

(* ===== HMI "HMI_RT_1" =====
system functions are stored by id; their names below are inferred from use

text list "Send Code Descriptions Short": 0 'SEND SUCCESSFUL'; 28672 'NO JOB'; 28673 'DATA ACCESSED DURING JOB'; 28674 'JOB PROCESSING'; 32901 'MAX LENGTH EXCEEDED'; 32902 'INVALID ID OUT OF RANGE'; 32904 'LENGTH EXCEEDS DATA RANGE'; 32929 'NO CONNECTION'; 32947 'UDP CONNECTION'; 32963 'CONNECTION BUSY'; 32964 'REQUEST DURING PARAM ASSIGNMENT'; 32965 'PARTNER TERMINATED CONNECTION'; 32966 'PARTNER UNAVAILABLE'; 32967 'TIMEOUT'; 65535 'NOT CALLED'

text list "Connect Code Descriptions Short": 0 'CONNECTION SUCCESSFUL'; 28672 'NO JOB'; 28673 'START JOB'; 28674 'PROCESSING JOB'; 32901 'ID INVALID: ALREADY IN USE'; 32902 'ID INVALID: OUT OF RANGE'; 32903 'MAX CONNECTIONS REACHED'; 32905 'NO CONNECTION DATA STORED'; 32922 'INVALID CONNECTION DATA'; 32923 'NO CONNECTION HARDWARE'; 32928 'GROUP ERROR'; 32929 'LOCAL PORT IN USE'; 32930 'REMOTE PORT IN USE'; 32931 'CONNECTION ALREADY ESTABLISHED'; 32932 'INVALID IP ADDRESS'; 32933 'DUPLICATE CONNECTION ID'; 32935 'DICONNECT REQUEST WHILE CONNECTING'; 32946 'CONNECT DATA IN LOAD MEMORY'; 32948 'ISO ON TCP VIOLATION'; 32949 'NON PASSIVE UDP CONNECTION REQUEST'; 32950 'INVALID CONNECTION TYPE'; 32951 'CONNECTION PARAMETER ERROR'; 32952 'DATA/PARAMETER MISMATCH'; 32963 'MAX CONNECTIONS EXCEEDED'; 32964 'FIREWALL'; 65535 'STATE: DISCONNECT'; 32966 'PARTNER UNAVAILABLE'

text list "Disconnect Code Descriptions Short": 0 'DISCONNECTION SUCCESSFUL'; 28672 'NO JOB'; 28673 'JOB STARTED'; 28674 'REQUEST DURING EXECUTION'; 32902 'ID INVALID: OUT OF RANGE'; 32931 'CONNECTION ALREADY TERMINATED'; 32964 'REQUEST DURING PARAM ASSIGNMENT'; 65535 'STATE: CONNECT'

text list "Text List Select": 0 ''; 1 ''; 2 ''; 3 ''

ScreenModuleEditorView "Connection_Status_Element" 392x110
   TextField "operation_label" at 0,0 size 110x110; Text 'S'
      Visibility <- "interface.operation_label_visible"
      Appearance <- "interface.operation_label_animate"
   TextField "done_status_indicator" at 110,0 size 94x27; Text 'DONE'
      Visibility <- "interface.done_status_indicator_visible"
      Appearance <- "interface.done_status_indicator_animate"
   TextField "busy_status_indicator" at 204,0 size 94x27; Text 'BUSY'
      Visibility <- "interface.busy_status_indicator_visible"
      Appearance <- "interface.busy_status_indicator_animate"
   TextField "error_status_indicator" at 298,0 size 94x27; Text 'ERROR'
      Visibility <- "interface.error_status_indicator_visible"
      Appearance <- "interface.error_status_indicator_animate"
   TextField "status_code_label" at 110,27 size 82x28; Text 'CODE:'
      Visibility <- "interface.status_code_label_visible"
      Appearance <- "interface.status_code_label_animate"
   IOField "status_code" at 192,27 size 200x28; FormatPattern ??????
      Appearance <- "interface.status_code_value_animate"
      Visibility <- "interface.status_code_value_visible"
      ProcessValue <- "interface.status_code_value"
   SymbolicIOField "status_description" at 110,55 size 282x55; TextOn '1'; TextOff '0'; TextList "Text List Select"
      Appearance <- "interface.status_code_description_animate"
      ProcessValue <- "operation_list_selector"
      Visibility <- "interface.status_code_description_visible"
   Button "operation_left" at 0,0 size 110x110; TextOff 'Text'
      on Press: function_b14e0dd5("interface.operation_button_actuate", 0)
      Visibility <- "interface.operation_button_visible"
      ObjectEnable <- "interface.operation_button_enable"
   Button "operation_top" at 110,0 size 282x55; TextOff 'Text'
      on Press: function_b14e0dd5("interface.operation_button_actuate", 0)
      Visibility <- "interface.operation_button_visible"
      ObjectEnable <- "interface.operation_button_enable"
   Button "show_status" at 110,55 size 282x55; TextOff 'Text'
      on Press: function_b14e0dd5("interface.show_status_code_description_button_actuate", 0)
      Visibility <- "interface.show_status_code_description_button_visible"
      ObjectEnable <- "interface.show_status_code_description_button_enable"
*)

(* ===== HMI "HMI_RT_1" =====
system functions are stored by id; their names below are inferred from use

text list "Connection Details Header": 0 'NO STATE'; 1 'DISCONNECTION STATUS'; 2 'CONNECTION STATUS'; 3 'SEND STATUS'

text list "Connect Code Descriptions Long": 0 'Connection successfully established.'; 28672 'No job processing active'; 28673 'Start job execution, establish connection.'; 28674 'Connection is being established (REQ irrelevant).'; 32901 'Connection ID (ID parameter) is already being used by a configured connection.'; 32902 'The ID parameter is outside the valid range.'; 32903 'Maximum number of connections reached; no additional connection possible'; 32905 'The CONNECT parameter does not point to a data block.'; 32922 'The structure at the CONNECT parameter is not supported on an integrated interface or the length is invalid or an incorrect "InterfaceID" is specified in the connection description (SDT).'; 32923 'The element InterfaceId within the TCON_xxx structure does not reference a hardware identifier of a CPU or CM/CP interface or has the value "0".'; 32928 'Group error for error codes W#16#80A1 and W#16#80A2.'; 32929 'The specified connection or the port is already being used.'; 32930 'Local or remote port is being used by the system.'; 32931 'Attempt being made to re-establish an existing connection.'; 32932 'IP address of the remote endpoint of the connection is invalid, in other words, it matches the IP address of the local partner.'; 32933 'Connection ID is already in use.'; 32935 'Communication error: You executed "TDISCON" before "TCON" had completed.'; 32946 'The CONNECT parameter points to a data block that was generated with the attribute "Only store in load memory".'; 32948 'ISO-on-TCP violation: local_tsap_id_len >= B#16#02 local_tsap_id[1] = B#16#E0 local_tsap_id_len >= B#16#03 local_tsap_id[1] is ASCII chr local_tsap_id[1] is ASCII cha and local_tsap_id_len >= B#16#03'; 32949 'Only passive connection establishment is permitted for connection type 13 = UDP.'; 32950 'Parameter assignment error at the connection_type parameter of the SDT TCON_Param.'; 32951 'Error in one of the following parameters of the data block for connection description: block_length, local_tsap_id_len, rem_subnet_id_len, rem_staddr_len, rem_tsap_id_len, next_staddr_len. Note: If you call TCON in TCP for the passive end, local_tsap_id_len must have the value 2 and rem_tsap_id_len the value 0.'; 32952 'Connection description of the structure element ID and the block parameter ID are not identical.'; 32963 'All connection resources are in use.'; 32964 'Temporary communication error: Firewall Pending Parameterization Pending Disconnect'; 65535 'In disconnect state.'; 32966 'The connection partner could not be reached.'